   'Open data source - Datenquelle öffnen
   conn.Open "Provider=MSDASQL;DSN="&Database_Name&"" 'DSN= name of the odbc-database - DSN= Name der ODBC-Datenbank
   
   'Error routine - Fehlerroutine
   If Err.Number <> 0 Then
   	bfde4b54-0db7-4817-8032-87127bf19bb9 "Error #" & Err.Number & " " & Err.Description
   	Err.Clear
   	Set conn = Nothing
   	Exit Sub
   End If
   
   
   'Create a database - Neue Datenbank erstellen
   SQL_Table = "CREATE DATABASE " & SmartTags("szDatabase")
   
   'Execute - Ausführen
   Set rst = conn.Execute(SQL_Table)
   
   'Error routine - Fehlerroutine
   If Err.Number <> 0 Then
   	bfde4b54-0db7-4817-8032-87127bf19bb9 "Error #" & Err.Number & " " & Err.Description
   	Err.Clear
   	'Close data source - Datenquelle schließen
   	conn.close
   	Set conn = Nothing
   	Set rst = Nothing
   	Exit Sub
   End If
   
   'Close data source - Datenquelle schließen
   conn.close
   
   Set conn = Nothing
   Set rst = Nothing

VB script "S01b_Delete_database"
   '////////////////////////////////////////////////////////////////
   ' en: The script deletes the indicated SQL database 
   ' de: Das Skript löscht die angegebene Datenbank
   ' Created: 19-07-2012
   ' Version: v1.0
   ' Author:  HH
   '////////////////////////////////////////////////////////////////
   
   'Declaration of local tags - Deklarartion von lokalen Variablen
   Dim conn, rst, SQL_Table
   
   On Error Resume Next
   
   Set conn = CreateObject("ADODB.Connection")
   Set rst = CreateObject("ADODB.Recordset")
   
   'Open data source - Datenquelle öffnen
   conn.Open "Provider=MSDASQL;DSN="&Database_Name&"" 'DSN= name of the odbc-database - DSN= Name der ODBC-Datenbank
   
   'Error routine - Fehlerroutine
   If Err.Number <> 0 Then
   	bfde4b54-0db7-4817-8032-87127bf19bb9 "Error #" & Err.Number & " " & Err.Description
   	Err.Clear
   	Set conn = Nothing
   	Exit Sub
   End If
   
   
   'Delete a database - Entfernt eine Datenbank
   SQL_Table = "DROP DATABASE " & SmartTags("szDatabase")
   
   'Execute - Ausführen
   Set rst = conn.Execute(SQL_Table)
   
   'Error routine - Fehlerroutine
   If Err.Number <> 0 Then
   	bfde4b54-0db7-4817-8032-87127bf19bb9 "Error #" & Err.Number & " " & Err.Description
   	Err.Clear
   	'Close data source - Datenquelle schließen
   	conn.close
   	Set conn = Nothing
   	Set rst = Nothing
   	Exit Sub
   End If
   
   'Close data source - Datenquelle schließen
   conn.close
   
   Set conn = Nothing
   Set rst = Nothing

VB script "S02_Create_new_table"
   '////////////////////////////////////////////////////////////////
   ' en: Creating a new table in the SQL database 
   ' de: Erstellen einer neuen Tablle in des SQL Datenbank
   ' Created: 19-07-2012
   ' Version: v1.0
   ' Author:  HH 
   '////////////////////////////////////////////////////////////////
   
   'Declaration of local tags - Deklaration von lokalen Variablen
   Dim conn, rst, SQL_Table
   
   On Error Resume Next
   
   Set conn = CreateObject("ADODB.Connection")
   Set rst = CreateObject("ADODB.Recordset")
   
   'Open data source - Datenquelle öffnen
   conn.Open "Provider=MSDASQL;Initial Catalog=" Lector620 ";DSN="&Database_Name&"" 'DSN= Name of the ODBC database - DSN= Name der ODBC-Datenbank
   
   'Error routine - Fehlerroutine
   If Err.Number <> 0 Then
   	bfde4b54-0db7-4817-8032-87127bf19bb9 "Error #" & Err.Number & " " & Err.Description
   	Err.Clear
   	Set conn = Nothing
   	Exit Sub
   End If
   
   
   'Create table - Tabelle erstellen
   'Definition of SQL table - Definition der SQL-Tabelle
   SQL_Table = "CREATE TABLE Crtne_Kode (Nr SMALLINT, " _
               & SmartTags("szName_1") & " CHAR(30), " & SmartTags("szName_2") & " SMALLINT, " _
               & SmartTags("szName_3") & " SMALLINT)"
   
   'Execute - Ausführen
   Set rst = conn.Execute(SQL_Table)
   
   'Error routine - Fehlerroutine 
   If Err.Number <> 0 Then
   	bfde4b54-0db7-4817-8032-87127bf19bb9 "Error #" & Err.Number & " " & Err.Description
   	Err.Clear
   	'Close data source - Datenquelle schließen
   	conn.close
   	Set conn = Nothing
   	Set rst = Nothing
   	Exit Sub
   End If
   
   'Close data source - Datenquelle schließen
   conn.close
   
   Set rst = Nothing
   Set conn = Nothing

VB script "S08_Copy_table"
   '////////////////////////////////////////////////////////////////
   ' en: Copy table containing the data records 
   ' de: Tabelle inklusive Datansatz kopieren
   ' Created: 19-07-2012
   ' Version: v1.0
   ' Author:  HH
   '////////////////////////////////////////////////////////////////
   
   'Declaration of local tags - Deklarartion von lokalen Variablen
   Dim conn, rst, SQL_Table
   
   On Error Resume Next
   
   Set conn = CreateObject("ADODB.Connection")
   Set rst = CreateObject("ADODB.Recordset")
   
   'Open data source - Datenquelle öffnen
   conn.Open "Provider=MSDASQL;Initial Catalog=" & SmartTags("szDatabase") & "; DSN="&Database_Name&"" 'DSN= Name der ODBC-Datenbank 'DSN= name of the odbc-database
   
   'Error routine - Fehlerroutine
   If Err.Number <> 0 Then
   	bfde4b54-0db7-4817-8032-87127bf19bb9 "Error #" & Err.Number & " " & Err.Description
   	Err.Clear
   	Set conn = Nothing
   	Exit Sub
   End If
   
   
   'Copying the SQL table - Kopieren der SQL Tabelle
   SQL_Table = " Select * Into " & SmartTags("szNewTableName") & " From " & SmartTags("szTableName")
   
   'Execute - Ausführen
   conn.execute(SQL_Table)
   
   'Error routine - Fehlerroutine
   If Err.Number <> 0 Then
   	bfde4b54-0db7-4817-8032-87127bf19bb9 "Error #" & Err.Number & " " & Err.Description
   	Err.Clear
   	'Close data source - Datenquelle schließen
   	conn.close
   	Set conn = Nothing
   	Set rst = Nothing
   	Exit Sub
   End If
   
   'Close data source - Datenquelle schließen
   conn.close
   
   Set rst = Nothing
   Set conn = Nothing

VB script "S09_Delete_table"
   '////////////////////////////////////////////////////////////////
   ' en: The script deletes the indicated table
   ' de: Das Skript löscht die angegebene Tabelle
   ' Created: 19-07-2012
   ' Version: v1.0
   ' Author:  HH
   '////////////////////////////////////////////////////////////////
   
   'Declarartion of local tags - Deklaration von lokalen Varaiblen
   Dim conn, rst, SQL_Table
   
   On Error Resume Next
   
   Set conn = CreateObject("ADODB.Connection")
   Set rst = CreateObject("ADODB.Recordset")
   
   'Open data source - Datenquelle öffnen
   conn.Open "Provider=MSDASQL;Initial Catalog=" & SmartTags("szDatabase") & ";DSN="&Database_Name&"" 'DSN= Name der ODBC-Datenbank 'DSN= name of the odbc-database
   
   'Error routine - Fehlerroutine
   If Err.Number <> 0 Then
   	bfde4b54-0db7-4817-8032-87127bf19bb9 "Error #" & Err.Number & " " & Err.Description
   	Err.Clear
   	Set conn = Nothing
   	Exit Sub
   End If
   
   
   'Delete table - Tabelle löschen
   SQL_Table = "DROP TABLE  "& SmartTags("szTableName")
   
   'Execute - Ausführen
   Set rst = conn.Execute(SQL_Table)
   
   'Error routine - Fehlerroutine
   If Err.Number <> 0 Then
   	bfde4b54-0db7-4817-8032-87127bf19bb9 "Error #" & Err.Number & " " & Err.Description
   	Err.Clear
   	'Close data source - Datenquelle schließen
   	conn.close
   	Set conn = Nothing
   	Set rst = Nothing
   	Exit Sub
   End If
   
   'Close data source - Datenquelle schließen
   conn.close
   
   Set rst = Nothing
   Set conn = Nothing

VB script "S04_Read_data_record_from_a_table"
   '////////////////////////////////////////////////////////////////
   ' en: The script reads the indicated data record
   ' de: Das Skript liest den angegebene Datensatz
   ' Created: 19-07-2012
   ' Version: v1.0
   ' Author:  HH 
   '////////////////////////////////////////////////////////////////
   
   'Declaration of local tags - Deklaration von lokalem Variablen
   Dim conn, rst, SQL_Table
   
   On Error Resume Next
   
   Set conn = CreateObject("ADODB.Connection")
   Set rst = CreateObject("ADODB.Recordset")
   
   'Open data source - Datenquelle öffnen
   conn.Open "Provider=MSDASQL;Initial Catalog=" & SmartTags("szDatabase") & ";DSN="&Database_Name&"" 'DSN= name of the odbc database - DSN= Name der ODBC-Datenbank
   
   'Error routine - Fehlerroutine
   If Err.Number <> 0 Then
   	bfde4b54-0db7-4817-8032-87127bf19bb9 "Error #" & Err.Number & " " & Err.Description
   	Err.Clear 
   	Set conn = Nothing
   	Exit Sub
   End If
   
   
   'Reads the data records of the SQL table
   'Select data record of the table - Datensatz der Tabelle auswählen
   SQL_Table = "SELECT * FROM " & SmartTags("szTableName") & " WHERE Nr = " & SmartTags("nDat_No")  '* = Alle Daten ' * = all data
   
   'Execute - Ausführen
   Set rst = conn.Execute(SQL_Table)
   
   'Error routine - Fehler Routine
   If Err.Number <> 0 Then
   	bfde4b54-0db7-4817-8032-87127bf19bb9 "Error #" & Err.Number & " " & Err.Description
   	Err.Clear
   	'Close data source - Datenquelle schließen
   	conn.close
   	Set conn = Nothing
   	Set rst = Nothing 
   	Exit Sub
   End If
   	
   If Not (rst.EOF And rst.BOF) Then 
   	'Vergleich ob End of File oder Begin of File ist, wenn nicht wird der Zeiger auf den ersten Eintrag zurueckgesetzt
   	'Compare if "End of File" or "Begin of File" exists, if not the pointer will be reset to the first entry
   	
   	rst.MoveFirst 'reset to 1st entry - auf 1. Eintrag zuruecksetzen 
   	
   	SmartTags("nDatNoTable") = rst.Fields(0).Value
   	SmartTags("nValue_1") = rst.Fields(1).Value
   	SmartTags("nValue_2") = rst.Fields(2).Value
   	SmartTags("nValue_3") = rst.Fields(3).Value 
   	SmartTags("szName_1") = rst.Fields(1).Name
   	SmartTags("szName_2") = rst.Fields(2).Name
   	SmartTags("szName_3") = rst.Fields(3).Name 
   	
   	rst.close 
   Else
   	bfde4b54-0db7-4817-8032-87127bf19bb9 "Dat_No. is not available"
   End If
   
   'Close data source - Datenquelle schließen
   conn.close
   
   Set rst = Nothing
   Set conn = Nothing

VB script "S03_Write_data_record_into_a_table"
   '////////////////////////////////////////////////////////////////
   ' en: The script wirtes the indicated data record into a table
   ' de: Das Skript schreibt den angegebene Datensatz in eine Tabelle
   ' Created: 19-07-2012
   ' Version: v1.0
   ' Author:  HH 
   '////////////////////////////////////////////////////////////////
   
   'Declaration of local tags - Deklaration von lokalen Variablen
   Dim conn, rst, SQL_Table
   
   On Error Resume Next
   
   Set conn = CreateObject("ADODB.Connection")
   Set rst = CreateObject("ADODB.Recordset")
   
   'Open data source - Datenquelle öffnen
   conn.Open "Provider=MSDASQL;Initial Catalog=" & SmartTags("szDatabase") & ";DSN="&Database_Name&"" 'DSN= Name of the ODBC database - DSN= Name der ODBC-Datenbank
   
   'Error routine - Fehlerroutine
   If Err.Number <> 0 Then
   	bfde4b54-0db7-4817-8032-87127bf19bb9 "Error #" & Err.Number & " " & Err.Description
   	Err.Clear
   	Set conn = Nothing 
   	Exit Sub
   End If
   
   
   'Writes a data record into a table
   'Select data record of the table - Datensatz der Tabelle auswählen
   SQL_Table = "SELECT * FROM " & SmartTags("szTableName") & " WHERE Nr = " & SmartTags("nDat_No")  '* = Alle Daten '* = all data
   
   'Execute - Ausführen
   Set rst = conn.Execute(SQL_Table)
   
   'Error routine - Fehler Routine
   If Err.Number <> 0 Then
   	bfde4b54-0db7-4817-8032-87127bf19bb9 "Error #" & Err.Number & " " & Err.Description
   	Err.Clear
   	'Close data source - Datenquelle schließen
   	conn.close
   	Set conn = Nothing
   	Set rst = Nothing 
   	Exit Sub
   End If
   
   If Not (rst.EOF And rst.BOF) Then 
   	'Compare if "End of File" or "Begin of File" exists, if not the pointer will be reset to the first entry
   	'Vergleich ob "End of File" oder "Begin of File" ist, wenn nicht wird der Zeiger auf den Ersten Eintrag zurueckgesetzt
    	bfde4b54-0db7-4817-8032-87127bf19bb9 "Dat No. exists already!"
   	rst.close 
   Else
   	'Definition of data record - Definition des Datensatzes
   	SQL_Table = "INSERT INTO "& SmartTags("szTableName") & " VALUES ('" & SmartTags("nDat_No") & _
   	            "' , '" & SmartTags("nValue_1") & "' , '" & SmartTags("nValue_2") & _
   	            "' , '" & SmartTags("nValue_3") & "')"
   	'Insert the data reacord of the table - Datensatz in die Tabelle hinzufügen
   	Set rst = conn.Execute(SQL_Table)
   End If
   
   'Close data source - Datenquelle schließen
   conn.close
   
   Set rst = Nothing
   Set conn = Nothing

VB script "S05_Edit_data_record"
   '////////////////////////////////////////////////////////////////
   ' en: The script updates the indicated data record
   ' de: Das Skript ändert den angegebene Datensatz
   ' Created: 19-07-2012
   ' Version: v1.0
   ' Author:  HH 
   '////////////////////////////////////////////////////////////////
   
   'Declaration of local tags - Deklaration von lokalen Varaiblen
   Dim conn, rst, SQL_Table
   
   On Error Resume Next
   
   Set conn = CreateObject("ADODB.Connection")
   Set rst = CreateObject("ADODB.Recordset")
   
   'Open data source - Datenquelle öffnen
   conn.Open "Provider=MSDASQL;Initial Catalog=" & SmartTags("szDatabase") & ";DSN="&Database_Name&"" 'DSN= Name der ODBC-Datenbank 'DSN= name of the odbc-database
   
   'Error routine - Fehlerroutine
   If Err.Number <> 0 Then
   	bfde4b54-0db7-4817-8032-87127bf19bb9 "Error #" & Err.Number & " " & Err.Description
   	Err.Clear 
   	Set conn = Nothing
   	Exit Sub
   End If
   
   
   'Reads the data records of the SQL table
   'Select data record of the table - Datensatz der Tabelle auswählen
   SQL_Table = "SELECT * FROM " & SmartTags("szTableName") & " WHERE Nr = " & SmartTags("nDat_No")  '* = Alle Daten ' * = all data
   
   'Execute - Ausführen
   Set rst = conn.Execute(SQL_Table)
   
   'Error routine - Fehler Routine
   If Err.Number <> 0 Then
   	bfde4b54-0db7-4817-8032-87127bf19bb9 "Error #" & Err.Number & " " & Err.Description
   	Err.Clear
   	'Close data source - Datenquelle schließen
   	conn.close
   	Set conn = Nothing
   	Set rst = Nothing 
   	Exit Sub
   End If
   	
   If Not (rst.EOF And rst.BOF) Then 
   	'Compare if "End of File" or "Begin of File" exists, if not the pointer will be reset to the first entry
   	'Vergleich ob End of File oder Begin of File ist, wenn nicht wird der Zeiger auf den Ersten Eintrag zurueckgesetzt
   		
   	rst.MoveFirst 'reset to 1st entry - auf 1. Eintrag zuruecksetzen 
   	 
   	SmartTags("szName_1") = rst.Fields(1).Name
   	SmartTags("szName_2") = rst.Fields(2).Name
   	SmartTags("szName_3") = rst.Fields(3).Name 
   	
   	rst.close 
   Else
   	bfde4b54-0db7-4817-8032-87127bf19bb9 "Dat_No. is not available" 'Ausgabe im ALARM VIEW, ob kein Eintrag 'dispaly at ALARM View, if no entry
   End If
   
   'Definition of data record - Definition des Datensatzes
   SQL_Table = "UPDATE "& SmartTags("szTableName") & " Set " & SmartTags("szName_1") & " = '" & SmartTags("nValue_1") & "' , " & SmartTags("szName_2") & " = " & SmartTags("nValue_2") & " , " & SmartTags("szName_3") & " = " & SmartTags("nValue_3") & " WHERE Nr = " & SmartTags("nDat_No") 
   
   'Update data record - Datensatz updaten
   Set rst = conn.Execute(SQL_Table)
   
   'Moja koda Stefan M---------------------------------------------------------------
   
   'SQL_Table = "UPDATE "& SmartTags("szTableName") & " Set " & SmartTags("szName_1") & " = '" & SmartTags("Code_read_string") & "' , " & SmartTags("iCounter_Tag_kopija") & " = " & SmartTags("nValue_2") & " , " & SmartTags("szName_3") & " = " & SmartTags("nValue_3") & " WHERE Nr = " & SmartTags("1") 
   
   
   'Konec----------------------------------------------------------------------------
   
   'Error routine - Fehlerroutine
   If Err.Number <> 0 Then
   	bfde4b54-0db7-4817-8032-87127bf19bb9 "Error #" & Err.Number & " " & Err.Description
   	Err.Clear
   	'Close data source - Datenquelle schließen
   	conn.close
   	Set conn = Nothing
   	Set rst = Nothing
   	Exit Sub
   End If
   
   'Close datab source - Datenquelle schließen
   conn.close
   
   Set rst = Nothing
   Set conn = Nothing

VB script "S06_Delete_data_record"
   '////////////////////////////////////////////////////////////////
   ' en: Creating a new table in the SQL database 
   ' de: Erstellen einer neuen Tablle in der SQL Datenbank
   ' Created: 19-07-2012
   ' Version: v1.0
   ' Author:  HH 
   '////////////////////////////////////////////////////////////////
   
   'Declaration of local tags - Deklaration von lokalen Variablen
   Dim conn, rst, SQL_Table
   
   On Error Resume Next
   
   Set conn = CreateObject("ADODB.Connection")
   Set rst = CreateObject("ADODB.Recordset")
   
   'Open data source - Datenquelle öffnen
   conn.Open "Provider=MSDASQL;Initial Catalog=" & SmartTags("szDatabase") & ";DSN="&Database_Name&"" 'DSN= Name der ODBC-Datenbank 'DSN= name of the odbc-database
   
   'Error routine - Fehlerroutine
   If Err.Number <> 0 Then
   	bfde4b54-0db7-4817-8032-87127bf19bb9 "Error #" & Err.Number & " " & Err.Description
   	Err.Clear
   	Set conn = Nothing 
   	Exit Sub
   End If
   
   
   'Delete data record - Datensatz aus Tabelle löschen
   SQL_Table = "DELETE FROM " & SmartTags("szTableName") &" WHERE Nr = " & SmartTags("nDat_No")  
   
   'Execute - Ausführen
   Set rst = conn.Execute(SQL_Table)
   
   'Error routine - Fehlerroutine
   If Err.Number <> 0 Then
   	bfde4b54-0db7-4817-8032-87127bf19bb9 "Error #" & Err.Number & " " & Err.Description
   	Err.Clear
   	'Close data source - Datenquelle schließen
   	conn.close
   	Set conn = Nothing
   	Set rst = Nothing
   	Exit Sub
   End If
   
   bfde4b54-0db7-4817-8032-87127bf19bb9 "Data record was deleted"
   
   'Close data source - Datenquelle schließen
   conn.close
   
   Set rst = Nothing
   Set conn = Nothing

VB script "TempScript"
   'Declaration of local tags - Deklaration von lokalen Variablen
   Dim conn, rst, SQL_Table
   
   On Error Resume Next
   
   Set conn = CreateObject("ADODB.Connection")
   Set rst = CreateObject("ADODB.Recordset")
   
   'Open data source - Datenquelle öffnen
   conn.Open "Provider=MSDASQL;Initial Catalog=Lector620;DSN="&Database_Name&"" 'DSN= Name of the ODBC database - DSN= Name der ODBC-Datenbank
   
   'Error routine - Fehlerroutine
   If Err.Number <> 0 Then
   	bfde4b54-0db7-4817-8032-87127bf19bb9 "Error #" & Err.Number & " " & Err.Description
   	Err.Clear
   	Set conn = Nothing 
   	Exit Sub
   End If
   
   
   	'Definition of data record - Definition des Datensatzes
   	SQL_Table = "INSERT INTO Crtne_Kode VALUES ('1' , '0606494564646546546' , '5' , '2008-01-01 00:00:01')"
   	'Insert the data reacord of the table - Datensatz in die Tabelle hinzufügen
   	Set rst = conn.Execute(SQL_Table)
   	
   	'Definition of data record - Definition des Datensatzes
   	SQL_Table = "INSERT INTO Crtne_Kode VALUES ('2' , '12121213' , '8' , '2009-06-08 12:04:05')"
   	'Insert the data reacord of the table - Datensatz in die Tabelle hinzufügen
   	Set rst = conn.Execute(SQL_Table)	
   	
   	'Definition of data record - Definition des Datensatzes
   	SQL_Table = "INSERT INTO Crtne_Kode VALUES ('3' , '878787878787' , '7' , '2015-09-012 05:07:08')"
   	'Insert the data reacord of the table - Datensatz in die Tabelle hinzufügen
   	Set rst = conn.Execute(SQL_Table)	
   	
   	'Definition of data record - Definition des Datensatzes
   	SQL_Table = "INSERT INTO Crtne_Kode VALUES ('4' , '9494949494' , '11' , '2020-08-01 08:10:08')"
   	'Insert the data reacord of the table - Datensatz in die Tabelle hinzufügen
   	Set rst = conn.Execute(SQL_Table)
   	
   	'Definition of data record - Definition des Datensatzes
   	SQL_Table = "INSERT INTO Crtne_Kode VALUES ('5' , '123456789' , '44' , '2021-12-30 12:11:10')"
   	'Insert the data reacord of the table - Datensatz in die Tabelle hinzufügen
   	Set rst = conn.Execute(SQL_Table)
   	
   	'Definition of data record - Definition des Datensatzes
   	SQL_Table = "INSERT INTO Crtne_Kode VALUES ('6' , '0987654321' , '112' , '2011-03-03 03:03:03')"
   	'Insert the data reacord of the table - Datensatz in die Tabelle hinzufügen
   	Set rst = conn.Execute(SQL_Table)
   	
   	
   'Error routine - Fehlerroutine
   If Err.Number <> 0 Then
   	bfde4b54-0db7-4817-8032-87127bf19bb9 "Error #" & Err.Number & " " & Err.Description
   	Err.Clear
   	'Close data source - Datenquelle schließen
   	conn.close
   	Set conn = Nothing
   	Set rst = Nothing
   	Exit Sub
   End If
   
   'Close data source - Datenquelle schließen
   conn.close
   
   Set rst = Nothing
   Set conn = Nothing

VB script "Branje_Artiklov"
   'Declaration of local tags - Deklaration von lokalen Variablen
   Dim conn, rst, SQL_Table, i, tempID
   
   On Error Resume Next
   
   Set conn = CreateObject("ADODB.Connection")
   Set rst = CreateObject("ADODB.Recordset")
   
   'Open data source - Datenquelle öffnen
   conn.Open "Provider=MSDASQL;Initial Catalog=Lector620;DSN="&Database_Name&"" 'DSN= Name of the ODBC database - DSN= Name der ODBC-Datenbank
   
   'Error routine - Fehlerroutine
   If Err.Number <> 0 Then
   	bfde4b54-0db7-4817-8032-87127bf19bb9 "Error #" & Err.Number & " " & Err.Description
   	Err.Clear
   	Set conn = Nothing 
   	Exit Sub
   End If
   
   '''''''''''''''''''''''
   	SmartTags("nTab")=0
   '''''''''''''''''''''''	
   
   	'Definition of data record - Definition des Datensatzes
   	SQL_Table = "SELECT COUNT(ID) FROM Crtne_Kode_Artiklov" 'Komanda v SQL v obliki string-a
   	'Insert the data record of the table - Datensatz in die Tabelle hinzufügen
   	Set rst = conn.Execute(SQL_Table) 'Komanda iz string-a se izvede
   	
   	If (rst.Fields(0).Value < 6) Then 'Nastavi i
   		
   		i=rst.Fields(0).Value
   		
   		Else i=6
   		
   	End If
   		
   		
   	
   	
   	'Vpisujemo parametre v tabelo v RT aplikaciji
   	
   	SQL_Table = "SELECT * FROM Crtne_Kode_Artiklov ORDER BY ID OFFSET 0 ROWS FETCH NEXT 6 ROWS ONLY"
   	Set rst = conn.Execute(SQL_Table)
   		
   	For i=0 To (i-1)
   		SmartTags("ID")(i)=rst.Fields(0).Value
   		SmartTags("tempID_Tag")(i)= rst.Fields(0).Value
   		SmartTags("Ime_Artikla_" & i)=CStr(rst.Fields(1).Value)
   		
   		SmartTags("Serijska_Stevilka_" & i)=CStr(rst.Fields(2).Value)
   		
   		
   		'SmartTags("Stevilo_Branja")(i)=rst.Fields(3).Value
   		
   		
   		SmartTags("Cas_Poslednjega_Branja")(i)=rst.Fields(4).Value
   		rst.MoveNext
   	Next
   	
   	
   
   	'Moramo posebej presteti koliko instanci enega artikla obstaja istega ID-a
   	For i=0 To (i-1)
   	SQL_Table = "SELECT COUNT(ID) FROM Crtne_Kode WHERE ID="&SmartTags("tempID_Tag")(i) 'Komanda v SQL v obliki string-a
   	Set rst = conn.Execute(SQL_Table) 'Komanda iz string-a se izvede
   	SmartTags("Stevilo_Branja")(i)=rst.Fields(0).Value
   	
   	
   	Next
   	
   	bfde4b54-0db7-4817-8032-87127bf19bb9 "Prebrano"
   	
   'Error routine - Fehlerroutine
   If Err.Number <> 0 Then
   	bfde4b54-0db7-4817-8032-87127bf19bb9 "Error #" & Err.Number & " " & Err.Description
   	Err.Clear
   	'Close data source - Datenquelle schließen
   	conn.close
   	Set conn = Nothing
   	Set rst = Nothing
   	Exit Sub
   End If
   
   'Close data source - Datenquelle schließen
   conn.close
   
   Set rst = Nothing
   Set conn = Nothing

VB script "Scrolling_Up_Down_Artikli"
   'Declaration of local tags - Deklaration von lokalen Variablen
   Dim conn, rst, SQL_Table, i
   
   On Error Resume Next
   
   Set conn = CreateObject("ADODB.Connection")
   Set rst = CreateObject("ADODB.Recordset")
   
   'Open data source - Datenquelle öffnen
   conn.Open "Provider=MSDASQL;Initial Catalog=Lector620;DSN="&Database_Name&"" 'DSN= Name of the ODBC database - DSN= Name der ODBC-Datenbank
   
   'Error routine - Fehlerroutine
   If Err.Number <> 0 Then
   	bfde4b54-0db7-4817-8032-87127bf19bb9 "Error #" & Err.Number & " " & Err.Description
   	Err.Clear
   	Set conn = Nothing 
   	Exit Sub
   End If
   
   	'Definition of data record - Definition des Datensatzes
   	SQL_Table = "SELECT COUNT(ID) FROM Crtne_Kode_Artiklov"
   	'Insert the data reacord of the table - Datensatz in die Tabelle hinzufügen
   	Set rst = conn.Execute(SQL_Table)
   	
   	If (rst.Fields(0).Value < 6) Then 
   		
   		i=rst.Fields(0).Value
   		
   		Else i=6
   		
   	End If
   	
   	If (SmartTags("nTab") > (rst.Fields(0).Value-6)) Then 
   		SmartTags("nTab")=rst.Fields(0).Value-6
   	End If		
   	
   	If (SmartTags("nTab") < 0) Then 
   		SmartTags("nTab")=0
   	End If
   	
   		
   		
   		
   	'Definition of data record - Definition des Datensatzes
   	SQL_Table = "SELECT * FROM Crtne_Kode_Artiklov ORDER BY ID OFFSET " &SmartTags("nTab")& " ROWS FETCH NEXT 6 ROWS ONLY"
   	'Insert the data reacord of the table - Datensatz in die Tabelle hinzufügen
   	Set rst = conn.Execute(SQL_Table)
   	
   	For i=0 To (i-1)
   		SmartTags("ID")(i)=rst.Fields(0).Value
   		
   		SmartTags("tempID_Tag")(i)= rst.Fields(0).Value
   		
   		SmartTags("Ime_Artikla_" & i)=rst.Fields(1).Value
   		
   		SmartTags("Serijska_Stevilka_" & i)=rst.Fields(2).Value
   		
   		SmartTags("Cas_Poslednjega_Branja")(i)=rst.Fields(4).Value
   		
   		rst.MoveNext
   	Next
   	
   	
   
   	'Moramo posebej presteti koliko instanci enega artikla obstaja istega ID-a
   	For i=0 To (i-1)
   	SQL_Table = "SELECT COUNT(ID) FROM Crtne_Kode WHERE ID="&SmartTags("tempID_Tag")(i) 'Komanda v SQL v obliki string-a
   	Set rst = conn.Execute(SQL_Table) 'Komanda iz string-a se izvede
   	SmartTags("Stevilo_Branja")(i)=rst.Fields(0).Value
   	
   	
   	Next
   	
   	
   'Error routine - Fehlerroutine
   If Err.Number <> 0 Then
   	bfde4b54-0db7-4817-8032-87127bf19bb9 "Error #" & Err.Number & " " & Err.Description
   	Err.Clear
   	'Close data source - Datenquelle schließen
   	conn.close
   	Set conn = Nothing
   	Set rst = Nothing
   	Exit Sub
   End If
   
   'Close data source - Datenquelle schließen
   conn.close
   
   Set rst = Nothing
   Set conn = Nothing

VB script "Sprejem_Serijske_Stevilke_v_SQL"
   'Declaration of local tags - Deklaration von lokalen Variablen
   Dim conn, rst, SQL_Table, tempID
   
   On Error Resume Next
   
   Set conn = CreateObject("ADODB.Connection")
   Set rst = CreateObject("ADODB.Recordset")
   
   'Open data source - Datenquelle öffnen
   conn.Open "Provider=MSDASQL;Initial Catalog=Lector620;DSN="&Database_Name&"" 'DSN= Name of the ODBC database - DSN= Name der ODBC-Datenbank
   
   'Error routine - Fehlerroutine
   If Err.Number <> 0 Then
   	bfde4b54-0db7-4817-8032-87127bf19bb9 "Error #" & Err.Number & " " & Err.Description
   	Err.Clear
   	Set conn = Nothing 
   	Exit Sub
   End If
   
   'Zacetek kode
   
   
   
   	
   	If (SmartTags("PrebranaKoda")<>"") Then
   	
   		If (SmartTags("PrebranaKoda")="NoRead") Then
   			bfde4b54-0db7-4817-8032-87127bf19bb9 "Nic ni prebrano, preverite ce senzor vidi kodo"
   						
   			Else
   			'Definition of data record - Definition des Datensatzes
   			SQL_Table = "SELECT * FROM Crtne_Kode_Artiklov WHERE Serijska_Stevilka='"&SmartTags("PrebranaKoda")&"'"
   			'Insert the data reacord of the table - Datensatz in die Tabelle hinzufügen
   			Set rst = conn.Execute(SQL_Table)
   			tempID=rst.Fields(0).Value
   			SmartTags("Novi_Artikel_Koda_Artikla_Temp")=SmartTags("PrebranaKoda")
   		
   		
   				If (rst.EOF And rst.BOF) Then
   				'Ce ni najdo kodo v sistemu
   				
   			
   				bfde4b54-0db7-4817-8032-87127bf19bb9 "Ne obstaja trenutno"
   				SmartTags("Nova_Serijska_Stevilka_Prebrana_ALARM")=1
   				'SmartTags("Novi_Artikel_Koda_Artikla_Temp")=SmartTags("PrebranaKoda")
   				SmartTags("Prebrana_Koda_FLAG")=1
   		
   		
   		
   		
   			
   				Else
   
   						
   							bfde4b54-0db7-4817-8032-87127bf19bb9 "Obstaja"
   							'Ce najde kodo ze v sistemu
   							
   							
   							SmartTags("Nova_Serijska_Stevilka_Prebrana_ALARM")=0
   							'SmartTags("Novi_Artikel_Koda_Artikla_Temp")=SmartTags("PrebranaKoda")
   							SmartTags("Prebrana_Koda_FLAG")=0
   							
   							SQL_Table ="INSERT INTO Crtne_Kode (ID,Cas_Poslednjega_Branja,Stanje) VALUES ('"&tempID&"',GETDATE(),'SKENIRAN!')"
   							
   							
   							
   					
   							Set rst = conn.Execute(SQL_Table) 'Komanda iz string-a se izvede
   						
   						
   							
   							'SQL_Table = "INSERT INTO Crtne_Kode (Serijska_Stevilka,Stevilo_Branja,Cas_Poslednjega_Branja) VALUES ( tempID ,GETDATE(),'OK!')"
   							'Insert the data reacord of the table - Datensatz in die Tabelle hinzufügen
   							'Set rst = conn.Execute(SQL_Table)
   							bfde4b54-0db7-4817-8032-87127bf19bb9 "Koda je uspesno dodana ustreznem artiklu"
   							SmartTags("Prebrana_Koda_FLAG")=0
   							
   							Scrolling_Up_Down_Artikli("Database_ArchiveMessage")
   		End If
   	End If
   End If
   
   'Konec Kode
   	
   	'SmartTags("PrebranaKoda")=""
   	
   	
   'Error routine - Fehlerroutine
   If Err.Number <> 0 Then
   	bfde4b54-0db7-4817-8032-87127bf19bb9 "Error #" & Err.Number & " " & Err.Description
   	Err.Clear
   	'Close data source - Datenquelle schließen
   	conn.close
   	Set conn = Nothing
   	Set rst = Nothing
   	Exit Sub
   End If
   
   'Close data source - Datenquelle schließen
   conn.close
   
   Set rst = Nothing
   Set conn = Nothing

VB script "Random"
   'TESTIRANJE
   
   
   'Declaration of local tags - Deklaration von lokalen Variablen
   Dim conn, rst, SQL_Table,Obj,return,return2,Tag
   
   On Error Resume Next
   
   Set conn = CreateObject("ADODB.Connection")
   Set rst = CreateObject("ADODB.Recordset")
   
   'Open data source - Datenquelle öffnen
   conn.Open "Provider=MSDASQL;Initial Catalog=Lector620;DSN="&Database_Name&"" 'DSN= Name of the ODBC database - DSN= Name der ODBC-Datenbank
   
   'Error routine - Fehlerroutine
   If Err.Number <> 0 Then
   	bfde4b54-0db7-4817-8032-87127bf19bb9 "Error #" & Err.Number & " " & Err.Description
   	Err.Clear
   	Set conn = Nothing 
   	Exit Sub
   End If
   
   
   
   	'Definition of data record - Definition des Datensatzes
   	'SQL_Table = "INSERT INTO Crtne_Kode_Artiklov (Serijska_Stevilka,Stevilo_Branja,Cas_Poslednjega_Branja) VALUES ('"&SmartTags("PrebranaKoda")&"','1',GETDATE())"
   	SQL_Table =	"INSERT INTO Crtne_Kode_Artiklov (Ime_Artikla,Serijska_Stevilka,Stevilo_Branja,Cas_Poslednjega_Branja) VALUES ('Mitsubishi_FX5UC AD','23456789987','1','2021-11-11 11:11:10.000')"
   	'Insert the data reacord of the table - Datensatz in die Tabelle hinzufügen
   	Set rst = conn.Execute(SQL_Table)
   	
   	
   
   
   	
   	
   'Error routine - Fehlerroutine
   If Err.Number <> 0 Then
   	bfde4b54-0db7-4817-8032-87127bf19bb9 "Error #" & Err.Number & " " & Err.Description
   	Err.Clear
   	'Close data source - Datenquelle schließen
   	conn.close
   	Set conn = Nothing
   	Set rst = Nothing
   	Exit Sub
   End If
   
   'Close data source - Datenquelle schließen
   conn.close
   
   Set rst = Nothing
   Set conn = Nothing

VB script "Iskanje_po_ID"
   'Declaration of local tags - Deklaration von lokalen Variablen
   Dim conn, rst, SQL_Table, i
   
   On Error Resume Next
   
   Set conn = CreateObject("ADODB.Connection")
   Set rst = CreateObject("ADODB.Recordset")
   
   'Open data source - Datenquelle öffnen
   conn.Open "Provider=MSDASQL;Initial Catalog=Lector620;DSN="&Database_Name&"" 'DSN= Name of the ODBC database - DSN= Name der ODBC-Datenbank
   
   'Error routine - Fehlerroutine
   If Err.Number <> 0 Then
   	bfde4b54-0db7-4817-8032-87127bf19bb9 "Error #" & Err.Number & " " & Err.Description
   	Err.Clear
   	Set conn = Nothing 
   	Exit Sub
   End If
   
   'Zacetek
   bfde4b54-0db7-4817-8032-87127bf19bb9 SmartTags("Iskanje_ID")
   	'Definition of data record - Definition des Datensatzes
   	SQL_Table = "SELECT COUNT(ID) FROM Crtne_Kode WHERE ID="&SmartTags("Iskanje_ID") 'Komanda v SQL v obliki string-a
   	'Insert the data record of the table - Datensatz in die Tabelle hinzufügen
   	Set rst = conn.Execute(SQL_Table) 'Komanda iz string-a se izvede
   	
   	 
   	
   	If (rst.Fields(0).Value < 6) Then 'Nastavi i
   		
   		i=rst.Fields(0).Value
   		
   		Else i=6
   		
   	End If
   		
   		
   	For i=0 To 5
   		SmartTags("ID")(i)=0
   		
   		SmartTags("Cas_Poslednjega_Branja")(i)=0
   		
   		SmartTags("Stanje_" & i)=""
   		
   		SmartTags("ID_Instance")(i)=0
   		
   	Next
   	
   	'Vpisujemo parametre v tabelo v RT aplikaciji
   	
   	SQL_Table = "SELECT * FROM Crtne_Kode WHERE ID="&SmartTags("Iskanje_ID")&" ORDER BY Cas_Poslednjega_Branja DESC OFFSET 0 ROWS FETCH NEXT 6 ROWS ONLY"
   	Set rst = conn.Execute(SQL_Table)
   		bfde4b54-0db7-4817-8032-87127bf19bb9 SmartTags("Iskanje_ID")
   	For i=0 To (i-1)
   		SmartTags("ID")(i)=rst.Fields(0).Value
   		
   		SmartTags("Cas_Poslednjega_Branja")(i)=rst.Fields(1).Value
   		
   		SmartTags("Stanje_" & i)=rst.Fields(2).Value
   		
   		SmartTags("ID_Instance")(i)=rst.Fields(3).Value
   		
   		rst.MoveNext
   	Next
   	
   
   'Konec
   
   
   
   
   
   'Error routine - Fehlerroutine
   If Err.Number <> 0 Then
   	bfde4b54-0db7-4817-8032-87127bf19bb9 "Error #" & Err.Number & " " & Err.Description
   	Err.Clear
   	'Close data source - Datenquelle schließen
   	conn.close
   	Set conn = Nothing
   	Set rst = Nothing
   	Exit Sub
   End If
   
   'Close data source - Datenquelle schließen
   conn.close
   
   Set rst = Nothing
   Set conn = Nothing

VB script "Iskanje_po_imenu_artikla"
   'Declaration of local tags - Deklaration von lokalen Variablen
   Dim conn, rst, SQL_Table, i, temp
   
   On Error Resume Next
   
   Set conn = CreateObject("ADODB.Connection")
   Set rst = CreateObject("ADODB.Recordset")
   
   'Open data source - Datenquelle öffnen
   conn.Open "Provider=MSDASQL;Initial Catalog=Lector620;DSN="&Database_Name&"" 'DSN= Name of the ODBC database - DSN= Name der ODBC-Datenbank
   
   'Error routine - Fehlerroutine
   If Err.Number <> 0 Then
   	bfde4b54-0db7-4817-8032-87127bf19bb9 "Error #" & Err.Number & " " & Err.Description
   	Err.Clear
   	Set conn = Nothing 
   	Exit Sub
   End If
   
   'Zacetek
   bfde4b54-0db7-4817-8032-87127bf19bb9 SmartTags("Iskanje_Instanci")
   	'Definition of data record - Definition des Datensatzes
   	SQL_Table = "SELECT COUNT(ID) FROM Crtne_Kode_Artiklov WHERE Ime_Artikla='"&SmartTags("Iskanje_Instanci")&"'" 'Komanda v SQL v obliki string-a
   	'Insert the data record of the table - Datensatz in die Tabelle hinzufügen
   	Set rst = conn.Execute(SQL_Table) 'Komanda iz string-a se izvede
   	
   	 
   	
   	If (rst.Fields(0).Value < 6) Then 'Nastavi i
   		
   		i=rst.Fields(0).Value
   		
   		Else i=6
   		
   	End If
   		
   		
   	For i=0 To 5
   		SmartTags("ID")(i)=0
   		
   		SmartTags("Cas_Poslednjega_Branja")(i)=0
   		
   		SmartTags("Stanje_" & i)=""
   		
   		SmartTags("ID_Instance")(i)=0
   
   	Next
   	
   	
   	'Vpisujemo parametre v tabelo v RT aplikaciji
   	
   	'Definition of data record - Definition des Datensatzes
   	SQL_Table = "SELECT ID FROM Crtne_Kode_Artiklov WHERE Ime_Artikla='"&SmartTags("Iskanje_Instanci")&"'" 'Komanda v SQL v obliki string-a
   	'Insert the data record of the table - Datensatz in die Tabelle hinzufügen
   	Set rst = conn.Execute(SQL_Table) 'Komanda iz string-a se izvede
   	
   	SmartTags("Iskanje_ID")=rst.Fields(0).Value
   	bfde4b54-0db7-4817-8032-87127bf19bb9 SmartTags("Iskanje_Instanci")
   	
   	SQL_Table = "SELECT * FROM Crtne_Kode WHERE ID="&SmartTags("Iskanje_ID")&" ORDER BY Cas_Poslednjega_Branja DESC OFFSET 0 ROWS FETCH NEXT 6 ROWS ONLY"
   	Set rst = conn.Execute(SQL_Table)
   		
   	For i=0 To (i-1)
   		SmartTags("ID")(i)=rst.Fields(0).Value
   		
   		SmartTags("Cas_Poslednjega_Branja")(i)=rst.Fields(1).Value
   		
   		SmartTags("Stanje_" & i)=rst.Fields(2).Value
   		
   		SmartTags("ID_Instance")(i)=rst.Fields(3).Value
   		
   		rst.MoveNext
   	Next
   	
   
   'Konec
   
   
   
   
   
   'Error routine - Fehlerroutine
   If Err.Number <> 0 Then
   	bfde4b54-0db7-4817-8032-87127bf19bb9 "Error #" & Err.Number & " " & Err.Description
   	Err.Clear
   	'Close data source - Datenquelle schließen
   	conn.close
   	Set conn = Nothing
   	Set rst = Nothing
   	Exit Sub
   End If
   
   'Close data source - Datenquelle schließen
   conn.close
   
   Set rst = Nothing
   Set conn = Nothing

VB script "Branje_Instanci_Artiklov"
   'Declaration of local tags - Deklaration von lokalen Variablen
   Dim conn, rst, SQL_Table, i, tempID
   
   On Error Resume Next
   
   Set conn = CreateObject("ADODB.Connection")
   Set rst = CreateObject("ADODB.Recordset")
   
   'Open data source - Datenquelle öffnen
   conn.Open "Provider=MSDASQL;Initial Catalog=Lector620;DSN="&Database_Name&"" 'DSN= Name of the ODBC database - DSN= Name der ODBC-Datenbank
   
   'Error routine - Fehlerroutine
   If Err.Number <> 0 Then
   	bfde4b54-0db7-4817-8032-87127bf19bb9 "Error #" & Err.Number & " " & Err.Description
   	Err.Clear
   	Set conn = Nothing 
   	Exit Sub
   End If
   
   '''''''''''''''''''''''
   	SmartTags("nTab")=0
   	SmartTags("Iskanje_ID")=0
   '''''''''''''''''''''''	
   	'Definition of data record - Definition des Datensatzes
   	SQL_Table = "SELECT COUNT(ID) FROM Crtne_Kode" 'Komanda v SQL v obliki string-a
   	'Insert the data record of the table - Datensatz in die Tabelle hinzufügen
   	Set rst = conn.Execute(SQL_Table) 'Komanda iz string-a se izvede
   	
   	If (rst.Fields(0).Value < 6) Then 'Nastavi i
   		
   		i=rst.Fields(0).Value
   		
   		Else i=6
   		
   	End If
   		
   		
   	
   	
   	'Vpisujemo parametre v tabelo v RT aplikaciji
   	
   	SQL_Table = "SELECT * FROM Crtne_Kode ORDER BY Cas_Poslednjega_Branja DESC OFFSET 0 ROWS FETCH NEXT 6 ROWS ONLY"
   	Set rst = conn.Execute(SQL_Table)
   		
   	For i=0 To (i-1)
   		SmartTags("ID")(i)=rst.Fields(0).Value
   		
   		SmartTags("Cas_Poslednjega_Branja")(i)=rst.Fields(1).Value	
   		
   		SmartTags("Stanje_" & i)=rst.Fields(2).Value
   		
   		SmartTags("ID_Instance")(i)=rst.Fields(3).Value
   		
   		rst.MoveNext
   	Next
   	
   	
   
   
   	
   	bfde4b54-0db7-4817-8032-87127bf19bb9 "Prebrano"
   	
   'Error routine - Fehlerroutine
   If Err.Number <> 0 Then
   	bfde4b54-0db7-4817-8032-87127bf19bb9 "Error #" & Err.Number & " " & Err.Description
   	Err.Clear
   	'Close data source - Datenquelle schließen
   	conn.close
   	Set conn = Nothing
   	Set rst = Nothing
   	Exit Sub
   End If
   
   'Close data source - Datenquelle schließen
   conn.close
   
   Set rst = Nothing
   Set conn = Nothing

VB script "Scrolling_Up_Down_Instanci"
   'Declaration of local tags - Deklaration von lokalen Variablen
   Dim conn, rst, SQL_Table, i,j
   
   On Error Resume Next
   
   Set conn = CreateObject("ADODB.Connection")
   Set rst = CreateObject("ADODB.Recordset")
   
   'Open data source - Datenquelle öffnen
   conn.Open "Provider=MSDASQL;Initial Catalog=Lector620;DSN="&Database_Name&"" 'DSN= Name of the ODBC database - DSN= Name der ODBC-Datenbank
   
   'Error routine - Fehlerroutine
   If Err.Number <> 0 Then
   	bfde4b54-0db7-4817-8032-87127bf19bb9 "Error #" & Err.Number & " " & Err.Description
   	Err.Clear
   	Set conn = Nothing 
   	Exit Sub
   End If
   
   
   	If (SmartTags("Iskanje_ID")<>0) Then
   
   	SQL_Table = "SELECT COUNT(ID) FROM Crtne_Kode WHERE ID="&SmartTags("Iskanje_ID")
   	
   	Else 
   		SQL_Table = "SELECT COUNT(ID) FROM Crtne_Kode"
   	
   	End If
   	Set rst = conn.Execute(SQL_Table)
   	
   	If (rst.Fields(0).Value < 6) Then 
   		
   		j=rst.Fields(0).Value
   		
   		Else j=6
   		
   	End If
   	
   		
   	If (SmartTags("nTab") > (rst.Fields(0).Value-6)) Then 
   		SmartTags("nTab")=rst.Fields(0).Value-6
   	End If	
   	
   	
   	If (SmartTags("nTab") < 0) Then 
   		SmartTags("nTab")=0
   	End If	
   		
   
   		
   	If (SmartTags("Iskanje_ID")<>0) Then	
   		
   	'Definition of data record - Definition des Datensatzes
   	SQL_Table = "SELECT * FROM Crtne_Kode WHERE ID="&SmartTags("Iskanje_ID")&" ORDER BY Cas_Poslednjega_Branja DESC OFFSET " &SmartTags("nTab")& " ROWS FETCH NEXT 6 ROWS ONLY"
   	'Insert the data reacord of the table - Datensatz in die Tabelle hinzufügen
   	
   	Else 
   		SQL_Table = "SELECT * FROM Crtne_Kode ORDER BY Cas_Poslednjega_Branja DESC OFFSET " &SmartTags("nTab")& " ROWS FETCH NEXT 6 ROWS ONLY"
   	
   	End If
   	
   	Set rst = conn.Execute(SQL_Table)
   	
   	bfde4b54-0db7-4817-8032-87127bf19bb9 ""&SmartTags("nTab")
   		
   	For i=0 To (j-1)
   		SmartTags("ID")(i)=rst.Fields(0).Value
   		
   		SmartTags("Cas_Poslednjega_Branja")(i)=rst.Fields(1).Value	
   		
   		SmartTags("Stanje_" & i)=rst.Fields(2).Value
   		
   		SmartTags("ID_Instance")(i)=rst.Fields(3).Value
   
   		rst.MoveNext
   	Next
   	
   
   
   
   	
   	
   'Error routine - Fehlerroutine
   If Err.Number <> 0 Then
   	bfde4b54-0db7-4817-8032-87127bf19bb9 "Error #" & Err.Number & " " & Err.Description
   	Err.Clear
   	'Close data source - Datenquelle schließen
   	conn.close
   	Set conn = Nothing
   	Set rst = Nothing
   	Exit Sub
   End If
   
   'Close data source - Datenquelle schließen
   conn.close
   
   Set rst = Nothing
   Set conn = Nothing

VB script "Sprejem_Serijske_Stevilke_v_SQL_Nova_Stevilka"
   'Declaration of local tags - Deklaration von lokalen Variablen
   Dim conn, rst, SQL_Table, tempID
   
   On Error Resume Next
   
   Set conn = CreateObject("ADODB.Connection")
   Set rst = CreateObject("ADODB.Recordset")
   
   'Open data source - Datenquelle öffnen
   conn.Open "Provider=MSDASQL;Initial Catalog=Lector620;DSN="&Database_Name&"" 'DSN= Name of the ODBC database - DSN= Name der ODBC-Datenbank
   
   'Error routine - Fehlerroutine
   If Err.Number <> 0 Then
   	bfde4b54-0db7-4817-8032-87127bf19bb9 "Error #" & Err.Number & " " & Err.Description
   	Err.Clear
   	Set conn = Nothing 
   	Exit Sub
   End If
   
   'Zacetek kode
   
   	 
   	'Definition of data record - Definition des Datensatzes
   	SQL_Table = "SELECT * FROM Crtne_Kode_Artiklov WHERE Serijska_Stevilka='"&SmartTags("PrebranaKoda")&"'"
   	'Insert the data reacord of the table - Datensatz in die Tabelle hinzufügen
   	Set rst = conn.Execute(SQL_Table)
       bfde4b54-0db7-4817-8032-87127bf19bb9 "vajda bela jakojako voli pavlakicu"
   	
   	If (rst.EOF And rst.BOF) Then
   		'Ce ni najdo kodo v sistemu
   		
   		
   			bfde4b54-0db7-4817-8032-87127bf19bb9 "Kreiranje novega artikla v poteku"
   			'If (SmartTags("Prebrana_Koda_FLAG")=1) Then
   				
   				'If (SmartTags("Novi_Artikel_Ime_Artikla_Temp")<>"") And (SmartTags("Novi_Artikel_Koda_Artikla_Temp") <> "") Then
   			
   			
   			'Vpisovanje tabela
   			SQL_Table = "INSERT INTO Crtne_Kode_Artiklov (Ime_Artikla,Serijska_Stevilka,Stevilo_Branja,Cas_Poslednjega_Branja) VALUES (  '"&SmartTags("Novi_Artikel_Ime_Artikla_Temp")&"','"&SmartTags("Novi_Artikel_Koda_Artikla_Temp")&"','1',GETDATE())"
   			Set rst = conn.Execute(SQL_Table)
   			
   			SQL_Table = "SELECT ID FROM Crtne_Kode_Artiklov WHERE Serijska_Stevilka='"&SmartTags("Novi_Artikel_Koda_Artikla_Temp")&"'"
   			'Insert the data reacord of the table - Datensatz in die Tabelle hinzufügen
   			Set rst = conn.Execute(SQL_Table)
   			
   			SmartTags("Novi_Artikel_ID_Artikla_Temp")=rst.Fields(0).Value
   			
   			
   			SQL_Table = "INSERT INTO Crtne_Kode (ID,Stanje,Cas_Poslednjega_Branja) VALUES ('"&SmartTags("Novi_Artikel_ID_Artikla_Temp")&"','SKENIRAN!',GETDATE())"
   			Set rst = conn.Execute(SQL_Table)
   			bfde4b54-0db7-4817-8032-87127bf19bb9 "uspelo3"
   			'
   			bfde4b54-0db7-4817-8032-87127bf19bb9 "Kreiranje novega artikla je bilo uspesno"
   				'Else
   					'ShowSystemAlarm "Parametri so nepravilno izpolnjeni"
   			
   			'End If
   		'End If
   	Else
   		'Ce najde kodo ze v sistemu
   			SmartTags("Novi_Artikel_ID_Artikla_Temp")=""
   			bfde4b54-0db7-4817-8032-87127bf19bb9 "Nikaj"
   			
   	End If
   
   
   'Konec Kode
   	
   	
   	
   	
   'Error routine - Fehlerroutine
   If Err.Number <> 0 Then
   	bfde4b54-0db7-4817-8032-87127bf19bb9 "Error #" & Err.Number & " " & Err.Description
   	Err.Clear
   	'Close data source - Datenquelle schließen
   	conn.close
   	Set conn = Nothing
   	Set rst = Nothing
   	Exit Sub
   End If
   
   'Close data source - Datenquelle schließen
   conn.close
   
   Set rst = Nothing
   Set conn = Nothing

VB script "Update_Stanja"
   'Declaration of local tags - Deklaration von lokalen Variablen
   Dim conn, rst, SQL_Table, tempStanjeidx
   
   On Error Resume Next
   
   Set conn = CreateObject("ADODB.Connection")
   Set rst = CreateObject("ADODB.Recordset")
   
   'Open data source - Datenquelle öffnen
   conn.Open "Provider=MSDASQL;Initial Catalog=Lector620;DSN="&Database_Name&"" 'DSN= Name of the ODBC database - DSN= Name der ODBC-Datenbank
   
   'Error routine - Fehlerroutine
   If Err.Number <> 0 Then
   	bfde4b54-0db7-4817-8032-87127bf19bb9 "Error #" & Err.Number & " " & Err.Description
   	Err.Clear
   	Set conn = Nothing 
   	Exit Sub
   End If
   
   'Zacetek
   
   	tempStanjeidx=SmartTags("Stanje_Update_Select")
   	SQL_Table = "SELECT Stanje FROM Crtne_Kode WHERE ID_Instance="&SmartTags("ID_Instance")(tempStanjeidx) 'Komanda v SQL v obliki string-a
   	Set rst = conn.Execute(SQL_Table) 'Komanda iz string-a se izvede
   	
   	 
   
   		If (rst.EOF And rst.BOF) Then
   			bfde4b54-0db7-4817-8032-87127bf19bb9 "Stef1"
   			bfde4b54-0db7-4817-8032-87127bf19bb9 "Napaka v posodabljanju stanja"
   		
   		Else
   			bfde4b54-0db7-4817-8032-87127bf19bb9 "Stef2"			
   			SQL_Table = "UPDATE Crtne_Kode SET Stanje='"&SmartTags("Stanje_"&tempStanjeidx)&"' WHERE ID_Instance="&SmartTags("ID_Instance")(tempStanjeidx)
   			Set rst = conn.Execute(SQL_Table) 'Komanda iz string-a se izvede		
   		End If
   
   	
   	
   	
   Scrolling_Up_Down_Instanci("Database_ArchiveMessage")
   'Konec
   
   
   
   
   
   'Error routine - Fehlerroutine
   If Err.Number <> 0 Then
   	bfde4b54-0db7-4817-8032-87127bf19bb9 "Error #" & Err.Number & " " & Err.Description
   	Err.Clear
   	'Close data source - Datenquelle schließen
   	conn.close
   	Set conn = Nothing
   	Set rst = Nothing
   	Exit Sub
   End If
   
   'Close data source - Datenquelle schließen
   conn.close
   
   Set rst = Nothing
   Set conn = Nothing

VB script "RT_Startup_Setup"
   If (SmartTags("Startup_Setup")=0) Then
   
   
   
   SmartTags("PrebranaKoda")=""
   
   
   
   
   
   SmartTags("Startup_Setup")=1
   End If

VB script "Posodobi_Iskanje_po_ID"
   'Declaration of local tags - Deklaration von lokalen Variablen
   Dim conn, rst, SQL_Table, i
   
   On Error Resume Next
   
   Set conn = CreateObject("ADODB.Connection")
   Set rst = CreateObject("ADODB.Recordset")
   
   'Open data source - Datenquelle öffnen
   conn.Open "Provider=MSDASQL;Initial Catalog=Lector620;DSN="&Database_Name&"" 'DSN= Name of the ODBC database - DSN= Name der ODBC-Datenbank
   
   'Error routine - Fehlerroutine
   If Err.Number <> 0 Then
   	bfde4b54-0db7-4817-8032-87127bf19bb9 "Error #" & Err.Number & " " & Err.Description
   	Err.Clear
   	Set conn = Nothing 
   	Exit Sub
   End If
   
   'Zacetek
   
   	'Definition of data record - Definition des Datensatzes
   	SQL_Table = "SELECT * FROM Crtne_Kode_Artiklov WHERE ID="&SmartTags("Novi_Artikel_ID_Artikla_Temp") 'Komanda v SQL v obliki string-a
   	'Insert the data record of the table - Datensatz in die Tabelle hinzufügen
   	Set rst = conn.Execute(SQL_Table) 'Komanda iz string-a se izvede
   	
   	 
   	
   	If (rst.EOF And rst.BOF) Then
   		
   		bfde4b54-0db7-4817-8032-87127bf19bb9 "Artikel ne obstaja!"
   		
   	Else 
   		
   		SmartTags("Novi_Artikel_Ime_Artikla_Temp")=rst.Fields(1).Value		
   		
   		SmartTags("Novi_Artikel_Koda_Artikla_Temp")=rst.Fields(2).Value		
   				
   	End If
   
   
   'Konec
   
   
   
   
   
   'Error routine - Fehlerroutine
   If Err.Number <> 0 Then
   	bfde4b54-0db7-4817-8032-87127bf19bb9 "Error #" & Err.Number & " " & Err.Description
   	Err.Clear
   	'Close data source - Datenquelle schließen
   	conn.close
   	Set conn = Nothing
   	Set rst = Nothing
   	Exit Sub
   End If
   
   'Close data source - Datenquelle schließen
   conn.close
   
   Set rst = Nothing
   Set conn = Nothing

VB script "Posodobi_Artikel"
   'Declaration of local tags - Deklaration von lokalen Variablen
   Dim conn, rst, SQL_Table, i, tempIme, tempKoda
   
   On Error Resume Next
   
   Set conn = CreateObject("ADODB.Connection")
   Set rst = CreateObject("ADODB.Recordset")
   
   'Open data source - Datenquelle öffnen
   conn.Open "Provider=MSDASQL;Initial Catalog=Lector620;DSN="&Database_Name&"" 'DSN= Name of the ODBC database - DSN= Name der ODBC-Datenbank
   
   'Error routine - Fehlerroutine
   If Err.Number <> 0 Then
   	bfde4b54-0db7-4817-8032-87127bf19bb9 "Error #" & Err.Number & " " & Err.Description
   	Err.Clear
   	Set conn = Nothing 
   	Exit Sub
   End If
   
   'Zacetek
   
   	'Definition of data record - Definition des Datensatzes
   	SQL_Table = "SELECT * FROM Crtne_Kode_Artiklov WHERE ID="&SmartTags("Novi_Artikel_ID_Artikla_Temp") 'Komanda v SQL v obliki string-a
   	'Insert the data record of the table - Datensatz in die Tabelle hinzufügen
   	Set rst = conn.Execute(SQL_Table) 'Komanda iz string-a se izvede
   	
   	tempIme=CStr(SmartTags("Novi_Artikel_Ime_Artikla_Temp"))	
   		
   	tempKoda=CStr(SmartTags("Novi_Artikel_Koda_Artikla_Temp"))		
   	 
   	
   	If (rst.EOF And rst.BOF) Then
   		
   		bfde4b54-0db7-4817-8032-87127bf19bb9 "Artikel ne obstaja!"
   		
   	Else 
   		
   			SQL_Table = "UPDATE Crtne_Kode_Artiklov SET Ime_Artikla='"&tempIme&"', Serijska_Stevilka='"&tempKoda&"' WHERE ID="&SmartTags("Novi_Artikel_ID_Artikla_Temp")
   			Set rst = conn.Execute(SQL_Table) 'Komanda iz string-a se izvede		
   		bfde4b54-0db7-4817-8032-87127bf19bb9 "Koncano"		
   	End If
   		
   		
   	
   		
   	
   		
   
   'Konec
   
   
   
   
   
   'Error routine - Fehlerroutine
   If Err.Number <> 0 Then
   	bfde4b54-0db7-4817-8032-87127bf19bb9 "Error #" & Err.Number & " " & Err.Description
   	Err.Clear
   	'Close data source - Datenquelle schließen
   	conn.close
   	Set conn = Nothing
   	Set rst = Nothing
   	Exit Sub
   End If
   
   'Close data source - Datenquelle schließen
   conn.close
   
   Set rst = Nothing
   Set conn = Nothing

VB script "IZBRISI_Artikel"
   'Declaration of local tags - Deklaration von lokalen Variablen
   Dim conn, rst, SQL_Table, i, tempIme, tempKoda
   
   On Error Resume Next
   
   Set conn = CreateObject("ADODB.Connection")
   Set rst = CreateObject("ADODB.Recordset")
   
   'Open data source - Datenquelle öffnen
   conn.Open "Provider=MSDASQL;Initial Catalog=Lector620;DSN="&Database_Name&"" 'DSN= Name of the ODBC database - DSN= Name der ODBC-Datenbank
   
   'Error routine - Fehlerroutine
   If Err.Number <> 0 Then
   	bfde4b54-0db7-4817-8032-87127bf19bb9 "Error #" & Err.Number & " " & Err.Description
   	Err.Clear
   	Set conn = Nothing 
   	Exit Sub
   End If
   
   'Zacetek
   
   	'Definition of data record - Definition des Datensatzes
   	SQL_Table = "SELECT * FROM Crtne_Kode_Artiklov WHERE ID="&SmartTags("Novi_Artikel_ID_Artikla_Temp") 'Komanda v SQL v obliki string-a
   	'Insert the data record of the table - Datensatz in die Tabelle hinzufügen
   	Set rst = conn.Execute(SQL_Table) 'Komanda iz string-a se izvede
   	 
   	
   	If (rst.EOF And rst.BOF) Then
   		
   		bfde4b54-0db7-4817-8032-87127bf19bb9 "Artikel ne obstaja!"
   		
   	Else 
   		
   			SQL_Table = "DELETE FROM Crtne_Kode_Artiklov WHERE ID="&SmartTags("Novi_Artikel_ID_Artikla_Temp")
   			Set rst = conn.Execute(SQL_Table) 'Komanda iz string-a se izvede		
   			bfde4b54-0db7-4817-8032-87127bf19bb9 "Brisanje Koncano!"		
   	End If
   		
   		
   	
   		
   	
   		
   
   'Konec
   
   
   
   
   
   'Error routine - Fehlerroutine
   If Err.Number <> 0 Then
   	bfde4b54-0db7-4817-8032-87127bf19bb9 "Error #" & Err.Number & " " & Err.Description
   	Err.Clear
   	'Close data source - Datenquelle schließen
   	conn.close
   	Set conn = Nothing
   	Set rst = Nothing
   	Exit Sub
   End If
   
   'Close data source - Datenquelle schließen
   conn.close
   
   Set rst = Nothing
   Set conn = Nothing
*)